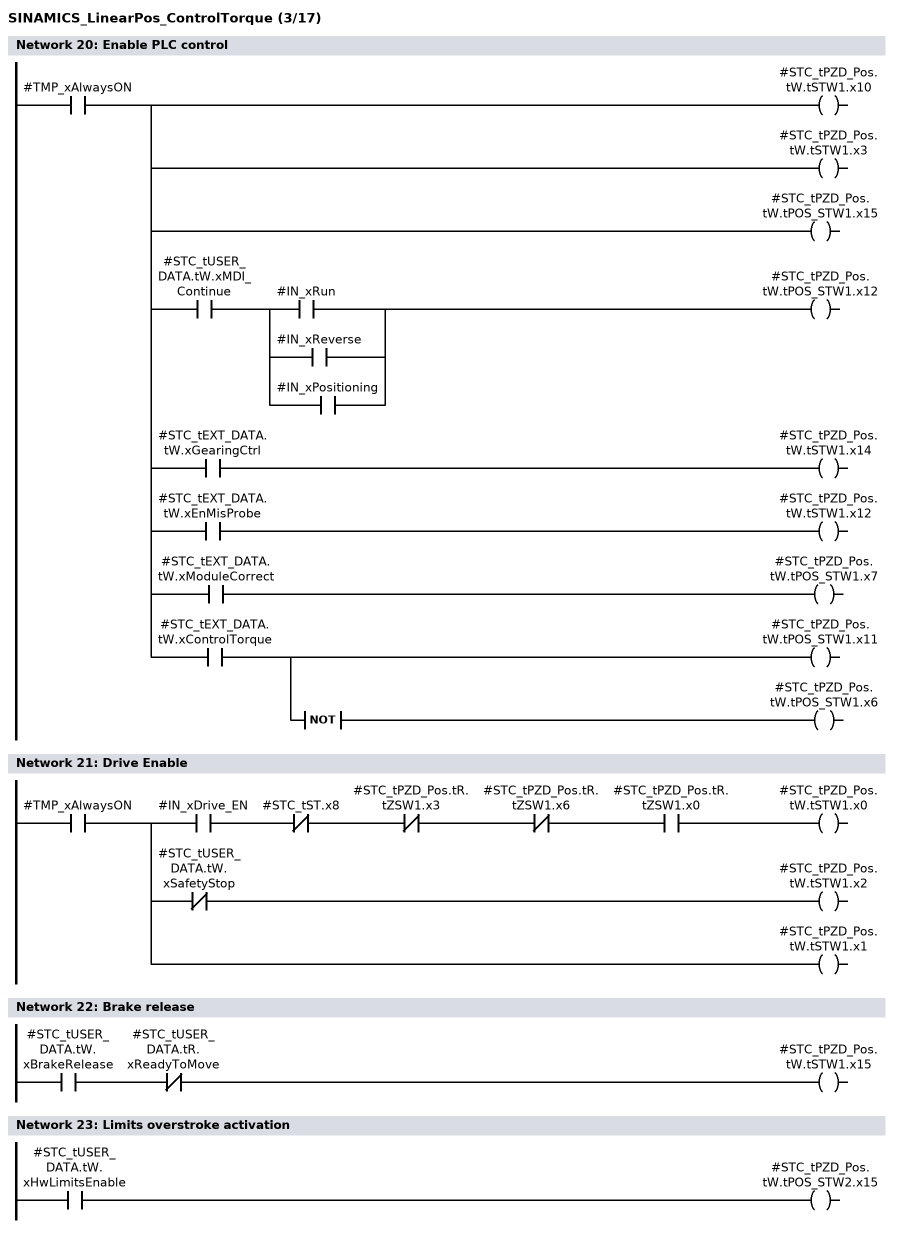
   RUNG wire#powerrail
      Contact( #TMP_xAlwaysON )
      wire#w1
      Coil( #STC_tPZD_Pos.tW.tSTW1.x10 )
   END_RUNG
   RUNG wire#w1
      Coil( #STC_tPZD_Pos.tW.tSTW1.x3 )
   END_RUNG
   RUNG wire#w1
      Coil( #STC_tPZD_Pos.tW.tPOS_STW1.x15 )
   END_RUNG
   RUNG wire#w1
      Contact( #STC_tUSER_DATA.tW.xMDI_Continue )
      wire#w2
      Contact( #IN_xRun )
      wire#w3
      Coil( #STC_tPZD_Pos.tW.tPOS_STW1.x12 )
   END_RUNG
   RUNG wire#w2
      Contact( #IN_xReverse )
   END_RUNG wire#w3
   RUNG wire#w2
      Contact( #IN_xPositioning )
   END_RUNG wire#w3
   RUNG wire#w1
      Contact( #STC_tEXT_DATA.tW.xGearingCtrl )
      Coil( #STC_tPZD_Pos.tW.tSTW1.x14 )
   END_RUNG
   RUNG wire#w1
      Contact( #STC_tEXT_DATA.tW.xEnMisProbe )
      Coil( #STC_tPZD_Pos.tW.tSTW1.x12 )
   END_RUNG
   RUNG wire#w1
      Contact( #STC_tEXT_DATA.tW.xModuleCorrect )
      Coil( #STC_tPZD_Pos.tW.tPOS_STW1.x7 )
   END_RUNG
   RUNG wire#w1
      Contact( #STC_tEXT_DATA.tW.xControlTorque )
      wire#w4
      Coil( #STC_tPZD_Pos.tW.tPOS_STW1.x11 )
   END_RUNG
   RUNG wire#w4
      Not()
      Coil( #STC_tPZD_Pos.tW.tPOS_STW1.x6 )
   END_RUNG
   // the same network as SCL:
   #STC_tPZD_Pos.tW.tSTW1.x10 := #TMP_xAlwaysON;
   #STC_tPZD_Pos.tW.tSTW1.x3 := #TMP_xAlwaysON;
   #STC_tPZD_Pos.tW.tPOS_STW1.x15 := #TMP_xAlwaysON;
   #STC_tPZD_Pos.tW.tPOS_STW1.x12 := #TMP_xAlwaysON AND #STC_tUSER_DATA.tW.xMDI_Continue AND (#IN_xRun OR #IN_xReverse OR #IN_xPositioning);
   #STC_tPZD_Pos.tW.tSTW1.x14 := #TMP_xAlwaysON AND #STC_tEXT_DATA.tW.xGearingCtrl;
   #STC_tPZD_Pos.tW.tSTW1.x12 := #TMP_xAlwaysON AND #STC_tEXT_DATA.tW.xEnMisProbe;
   #STC_tPZD_Pos.tW.tPOS_STW1.x7 := #TMP_xAlwaysON AND #STC_tEXT_DATA.tW.xModuleCorrect;
   #STC_tPZD_Pos.tW.tPOS_STW1.x11 := #TMP_xAlwaysON AND #STC_tEXT_DATA.tW.xControlTorque;
   #STC_tPZD_Pos.tW.tPOS_STW1.x6 := NOT #STC_tPZD_Pos.tW.tPOS_STW1.x11;
END_REGION

REGION Network 21: Drive Enable
   RUNG wire#powerrail
      Contact( #TMP_xAlwaysON )
      wire#w1
      Contact( #IN_xDrive_EN )
      I_Contact( #STC_tST.x8 )
      I_Contact( #STC_tPZD_Pos.tR.tZSW1.x3 )
      I_Contact( #STC_tPZD_Pos.tR.tZSW1.x6 )
      Contact( #STC_tPZD_Pos.tR.tZSW1.x0 )
      Coil( #STC_tPZD_Pos.tW.tSTW1.x0 )
   END_RUNG
   RUNG wire#w1
      I_Contact( #STC_tUSER_DATA.tW.xSafetyStop )
      Coil( #STC_tPZD_Pos.tW.tSTW1.x2 )
   END_RUNG
   RUNG wire#w1
      Coil( #STC_tPZD_Pos.tW.tSTW1.x1 )
   END_RUNG
   // the same network as SCL:
   #STC_tPZD_Pos.tW.tSTW1.x0 := #TMP_xAlwaysON AND #IN_xDrive_EN AND NOT #STC_tST.x8 AND NOT #STC_tPZD_Pos.tR.tZSW1.x3 AND NOT #STC_tPZD_Pos.tR.tZSW1.x6 AND #STC_tPZD_Pos.tR.tZSW1.x0;
   #STC_tPZD_Pos.tW.tSTW1.x2 := #TMP_xAlwaysON AND NOT #STC_tUSER_DATA.tW.xSafetyStop;
   #STC_tPZD_Pos.tW.tSTW1.x1 := #TMP_xAlwaysON;
END_REGION

REGION Network 22: Brake release
   RUNG wire#powerrail
      Contact( #STC_tUSER_DATA.tW.xBrakeRelease )
      I_Contact( #STC_tUSER_DATA.tR.xReadyToMove )
      Coil( #STC_tPZD_Pos.tW.tSTW1.x15 )
   END_RUNG
   // the same network as SCL:
   #STC_tPZD_Pos.tW.tSTW1.x15 := #STC_tUSER_DATA.tW.xBrakeRelease AND NOT #STC_tUSER_DATA.tR.xReadyToMove;
END_REGION

REGION Network 23: Limits overstroke activation
   RUNG wire#powerrail
      Contact( #STC_tUSER_DATA.tW.xHwLimitsEnable )
      Coil( #STC_tPZD_Pos.tW.tPOS_STW2.x15 )
   END_RUNG
   // the same network as SCL:
   #STC_tPZD_Pos.tW.tPOS_STW2.x15 := #STC_tUSER_DATA.tW.xHwLimitsEnable;
END_REGION

REGION Network 24: OS.Fly referencing active
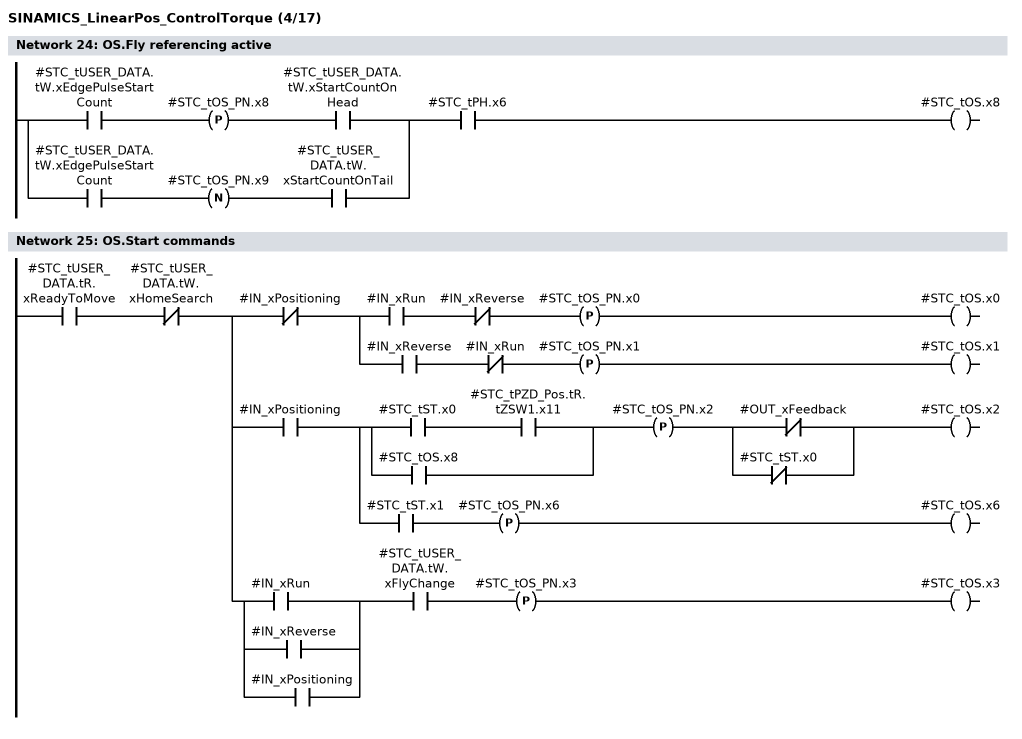
   RUNG wire#powerrail
      Contact( #STC_tUSER_DATA.tW.xEdgePulseStartCount )
      P_Trig( #STC_tOS_PN.x8 )
      Contact( #STC_tUSER_DATA.tW.xStartCountOnHead )
      wire#w1
      Contact( #STC_tPH.x6 )
      Coil( #STC_tOS.x8 )
   END_RUNG
   RUNG wire#powerrail
      Contact( #STC_tUSER_DATA.tW.xEdgePulseStartCount )
      N_Trig( #STC_tOS_PN.x9 )
      Contact( #STC_tUSER_DATA.tW.xStartCountOnTail )
   END_RUNG wire#w1
   // the same network as SCL:
   #_w1 := #STC_tUSER_DATA.tW.xEdgePulseStartCount AND NOT #STC_tOS_PN.x8;   // rising edge
   #STC_tOS_PN.x8 := #STC_tUSER_DATA.tW.xEdgePulseStartCount;
   #_w2 := NOT #STC_tUSER_DATA.tW.xEdgePulseStartCount AND #STC_tOS_PN.x9;   // falling edge
   #STC_tOS_PN.x9 := #STC_tUSER_DATA.tW.xEdgePulseStartCount;
   #STC_tOS.x8 := ((#_w1 AND #STC_tUSER_DATA.tW.xStartCountOnHead) OR (#_w2 AND #STC_tUSER_DATA.tW.xStartCountOnTail)) AND #STC_tPH.x6;
END_REGION

REGION Network 25: OS.Start commands
   RUNG wire#powerrail
      Contact( #STC_tUSER_DATA.tR.xReadyToMove )
      I_Contact( #STC_tUSER_DATA.tW.xHomeSearch )
      wire#w1
      I_Contact( #IN_xPositioning )
      wire#w2
      Contact( #IN_xRun )
      I_Contact( #IN_xReverse )
      P_Trig( #STC_tOS_PN.x0 )
      Coil( #STC_tOS.x0 )
   END_RUNG
   RUNG wire#w2
      Contact( #IN_xReverse )
      I_Contact( #IN_xRun )
      P_Trig( #STC_tOS_PN.x1 )
      Coil( #STC_tOS.x1 )
   END_RUNG
   RUNG wire#w1
      Contact( #IN_xPositioning )
      wire#w3
      Contact( #STC_tST.x0 )
      Contact( #STC_tPZD_Pos.tR.tZSW1.x11 )
      wire#w4
      P_Trig( #STC_tOS_PN.x2 )
      wire#w5
      I_Contact( #OUT_xFeedback )
      wire#w6
      Coil( #STC_tOS.x2 )
   END_RUNG
   RUNG wire#w3
      Contact( #STC_tOS.x8 )
   END_RUNG wire#w4
   RUNG wire#w5
      I_Contact( #STC_tST.x0 )
   END_RUNG wire#w6
   RUNG wire#w3
      Contact( #STC_tST.x1 )
      P_Trig( #STC_tOS_PN.x6 )
      Coil( #STC_tOS.x6 )
   END_RUNG
   RUNG wire#w1
      Contact( #IN_xRun )
      wire#w7
      Contact( #STC_tUSER_DATA.tW.xFlyChange )
      P_Trig( #STC_tOS_PN.x3 )
      Coil( #STC_tOS.x3 )
   END_RUNG
   RUNG wire#w1
      Contact( #IN_xReverse )
   END_RUNG wire#w7
   RUNG wire#w1
      Contact( #IN_xPositioning )
   END_RUNG wire#w7
   // the same network as SCL:
   #_w1 := #STC_tUSER_DATA.tR.xReadyToMove AND NOT #STC_tUSER_DATA.tW.xHomeSearch;
   #_w2 := #_w1 AND NOT #IN_xPositioning;
   #_w3 := #_w2 AND #IN_xRun AND NOT #IN_xReverse;
   #_w4 := #_w3 AND NOT #STC_tOS_PN.x0;   // rising edge
   #STC_tOS_PN.x0 := #_w3;
   #STC_tOS.x0 := #_w4;
   #_w5 := #_w2 AND #IN_xReverse AND NOT #IN_xRun;
   #_w6 := #_w5 AND NOT #STC_tOS_PN.x1;   // rising edge
   #STC_tOS_PN.x1 := #_w5;
   #STC_tOS.x1 := #_w6;
   #_w7 := #_w1 AND #IN_xPositioning;
   #_w8 := #_w7 AND ((#STC_tST.x0 AND #STC_tPZD_Pos.tR.tZSW1.x11) OR #STC_tOS.x8);
   #_w9 := #_w8 AND NOT #STC_tOS_PN.x2;   // rising edge
   #STC_tOS_PN.x2 := #_w8;
   #STC_tOS.x2 := #_w9 AND (NOT #OUT_xFeedback OR NOT #STC_tST.x0);
   #_w10 := #_w7 AND #STC_tST.x1;
   #_w11 := #_w10 AND NOT #STC_tOS_PN.x6;   // rising edge
   #STC_tOS_PN.x6 := #_w10;
   #STC_tOS.x6 := #_w11;
   #_w12 := #_w1 AND (#IN_xRun OR #IN_xReverse OR #IN_xPositioning) AND #STC_tUSER_DATA.tW.xFlyChange;
   #_w13 := #_w12 AND NOT #STC_tOS_PN.x3;   // rising edge
   #STC_tOS_PN.x3 := #_w12;
   #STC_tOS.x3 := #_w13;
END_REGION

REGION Network 26: Sending data copy
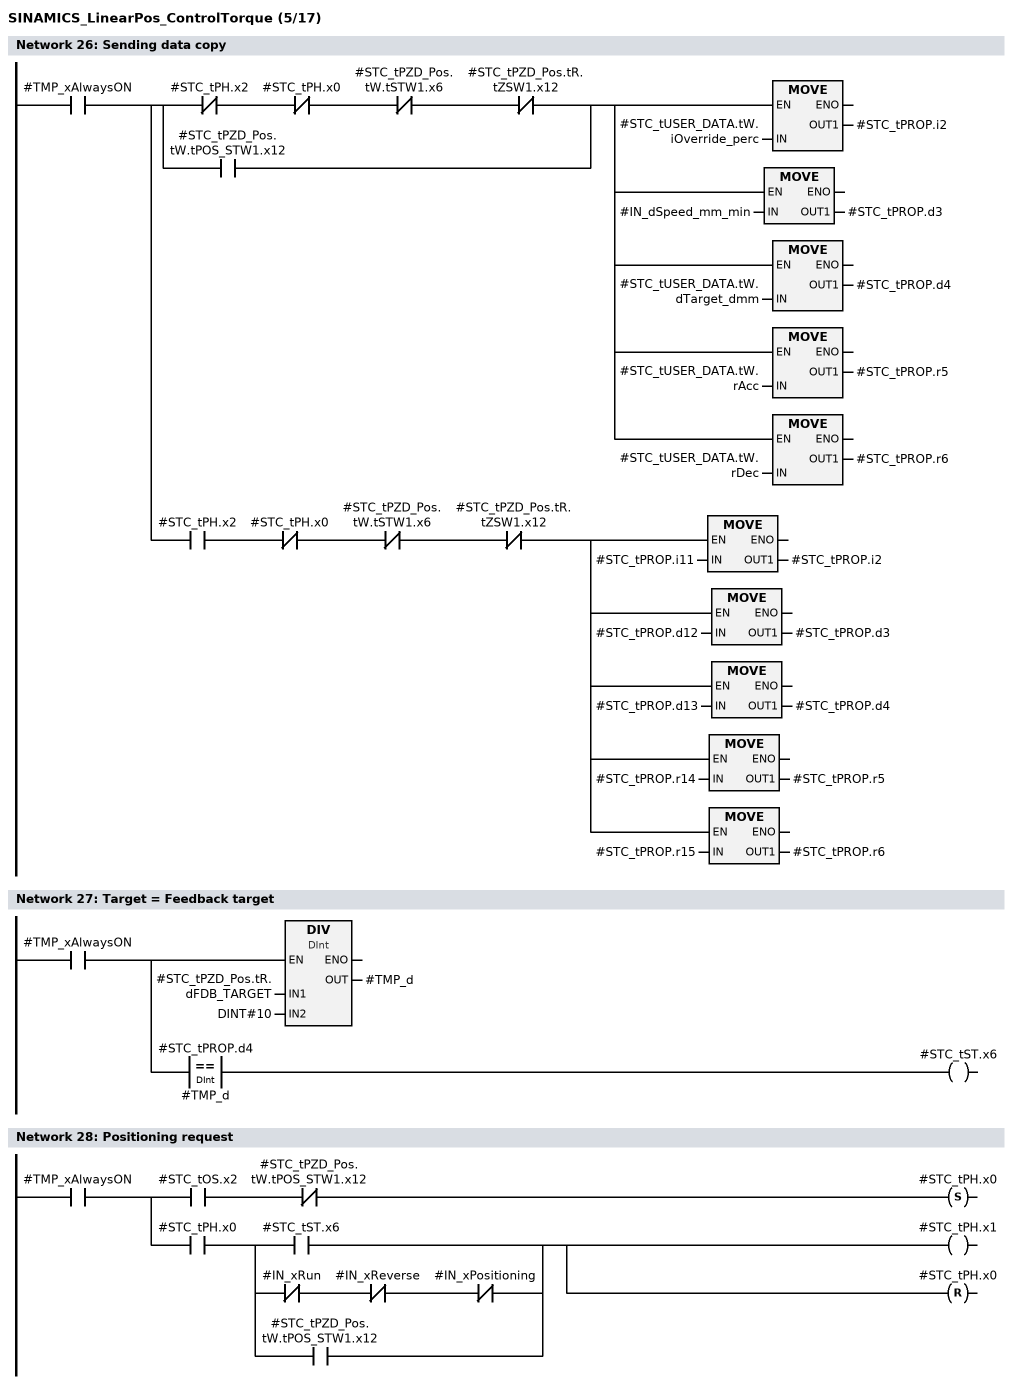
   RUNG wire#powerrail
      Contact( #TMP_xAlwaysON )
      wire#w1
      I_Contact( #STC_tPH.x2 )
      I_Contact( #STC_tPH.x0 )
      I_Contact( #STC_tPZD_Pos.tW.tSTW1.x6 )
      I_Contact( #STC_tPZD_Pos.tR.tZSW1.x12 )
      wire#w2
      { S7_GenerateENO := "TRUE" } Move(in := #STC_tUSER_DATA.tW.iOverride_perc, out1 => #STC_tPROP.i2)
   END_RUNG
   RUNG wire#w1
      Contact( #STC_tPZD_Pos.tW.tPOS_STW1.x12 )
   END_RUNG wire#w2
   RUNG wire#w2
      { S7_GenerateENO := "TRUE" } Move(in := #IN_dSpeed_mm_min, out1 => #STC_tPROP.d3)
   END_RUNG
   RUNG wire#w2
      { S7_GenerateENO := "TRUE" } Move(in := #STC_tUSER_DATA.tW.dTarget_dmm, out1 => #STC_tPROP.d4)
   END_RUNG
   RUNG wire#w2
      { S7_GenerateENO := "TRUE" } Move(in := #STC_tUSER_DATA.tW.rAcc, out1 => #STC_tPROP.r5)
   END_RUNG
   RUNG wire#w2
      { S7_GenerateENO := "TRUE" } Move(in := #STC_tUSER_DATA.tW.rDec, out1 => #STC_tPROP.r6)
   END_RUNG
   RUNG wire#w1
      Contact( #STC_tPH.x2 )
      I_Contact( #STC_tPH.x0 )
      I_Contact( #STC_tPZD_Pos.tW.tSTW1.x6 )
      I_Contact( #STC_tPZD_Pos.tR.tZSW1.x12 )
      wire#w3
      { S7_GenerateENO := "TRUE" } Move(in := #STC_tPROP.i11, out1 => #STC_tPROP.i2)
   END_RUNG
   RUNG wire#w3
      { S7_GenerateENO := "TRUE" } Move(in := #STC_tPROP.d12, out1 => #STC_tPROP.d3)
   END_RUNG
   RUNG wire#w3
      { S7_GenerateENO := "TRUE" } Move(in := #STC_tPROP.d13, out1 => #STC_tPROP.d4)
   END_RUNG
   RUNG wire#w3
      { S7_GenerateENO := "TRUE" } Move(in := #STC_tPROP.r14, out1 => #STC_tPROP.r5)
   END_RUNG
   RUNG wire#w3
      { S7_GenerateENO := "TRUE" } Move(in := #STC_tPROP.r15, out1 => #STC_tPROP.r6)
   END_RUNG
   // the same network as SCL:
   IF #TMP_xAlwaysON AND ((NOT #STC_tPH.x2 AND NOT #STC_tPH.x0 AND NOT #STC_tPZD_Pos.tW.tSTW1.x6 AND NOT #STC_tPZD_Pos.tR.tZSW1.x12) OR #STC_tPZD_Pos.tW.tPOS_STW1.x12) THEN
       #STC_tPROP.i2 := #STC_tUSER_DATA.tW.iOverride_perc;
       #STC_tPROP.d3 := #IN_dSpeed_mm_min;
       #STC_tPROP.d4 := #STC_tUSER_DATA.tW.dTarget_dmm;
       #STC_tPROP.r5 := #STC_tUSER_DATA.tW.rAcc;
       #STC_tPROP.r6 := #STC_tUSER_DATA.tW.rDec;
   END_IF;
   IF #TMP_xAlwaysON AND #STC_tPH.x2 AND NOT #STC_tPH.x0 AND NOT #STC_tPZD_Pos.tW.tSTW1.x6 AND NOT #STC_tPZD_Pos.tR.tZSW1.x12 THEN
       #STC_tPROP.i2 := #STC_tPROP.i11;
       #STC_tPROP.d3 := #STC_tPROP.d12;
       #STC_tPROP.d4 := #STC_tPROP.d13;
       #STC_tPROP.r5 := #STC_tPROP.r14;
       #STC_tPROP.r6 := #STC_tPROP.r15;
   END_IF;
END_REGION

REGION Network 27: Target = Feedback target
   RUNG wire#powerrail
      Contact( #TMP_xAlwaysON )
      wire#w1
      { S7_Templates := "SrcType := DInt"; S7_GenerateENO := "TRUE" } Div(in1 := #STC_tPZD_Pos.tR.dFDB_TARGET, in2 := DINT#10, out => #TMP_d)
   END_RUNG
   RUNG wire#w1
      { S7_Templates := "SrcType := DInt" } EQ_Contact(in1 := #STC_tPROP.d4, in2 := #TMP_d)
      Coil( #STC_tST.x6 )
   END_RUNG
   // the same network as SCL:
   IF #TMP_xAlwaysON THEN #TMP_d := #STC_tPZD_Pos.tR.dFDB_TARGET / DINT#10; END_IF;
   #STC_tST.x6 := #TMP_xAlwaysON AND (#STC_tPROP.d4 = #TMP_d);
END_REGION

REGION Network 28: Positioning request
   RUNG wire#powerrail
      Contact( #TMP_xAlwaysON )
      wire#w1
      Contact( #STC_tOS.x2 )
      I_Contact( #STC_tPZD_Pos.tW.tPOS_STW1.x12 )
      S_Coil( #STC_tPH.x0 )
   END_RUNG
   RUNG wire#w1
      Contact( #STC_tPH.x0 )
      wire#w2
      Contact( #STC_tST.x6 )
      wire#w3
      Coil( #STC_tPH.x1 )
   END_RUNG
   RUNG wire#w2
      I_Contact( #IN_xRun )
      I_Contact( #IN_xReverse )
      I_Contact( #IN_xPositioning )
   END_RUNG wire#w3
   RUNG wire#w2
      Contact( #STC_tPZD_Pos.tW.tPOS_STW1.x12 )
   END_RUNG wire#w3
   RUNG wire#w3
      R_Coil( #STC_tPH.x0 )
   END_RUNG
   // the same network as SCL:
   IF #TMP_xAlwaysON AND #STC_tOS.x2 AND NOT #STC_tPZD_Pos.tW.tPOS_STW1.x12 THEN #STC_tPH.x0 := TRUE; END_IF;
   #STC_tPH.x1 := #TMP_xAlwaysON AND #STC_tPH.x0 AND (#STC_tST.x6 OR (NOT #IN_xRun AND NOT #IN_xReverse AND NOT #IN_xPositioning) OR #STC_tPZD_Pos.tW.tPOS_STW1.x12);
   IF #STC_tPH.x1 THEN #STC_tPH.x0 := FALSE; END_IF;
END_REGION

REGION Network 29: Fly change request
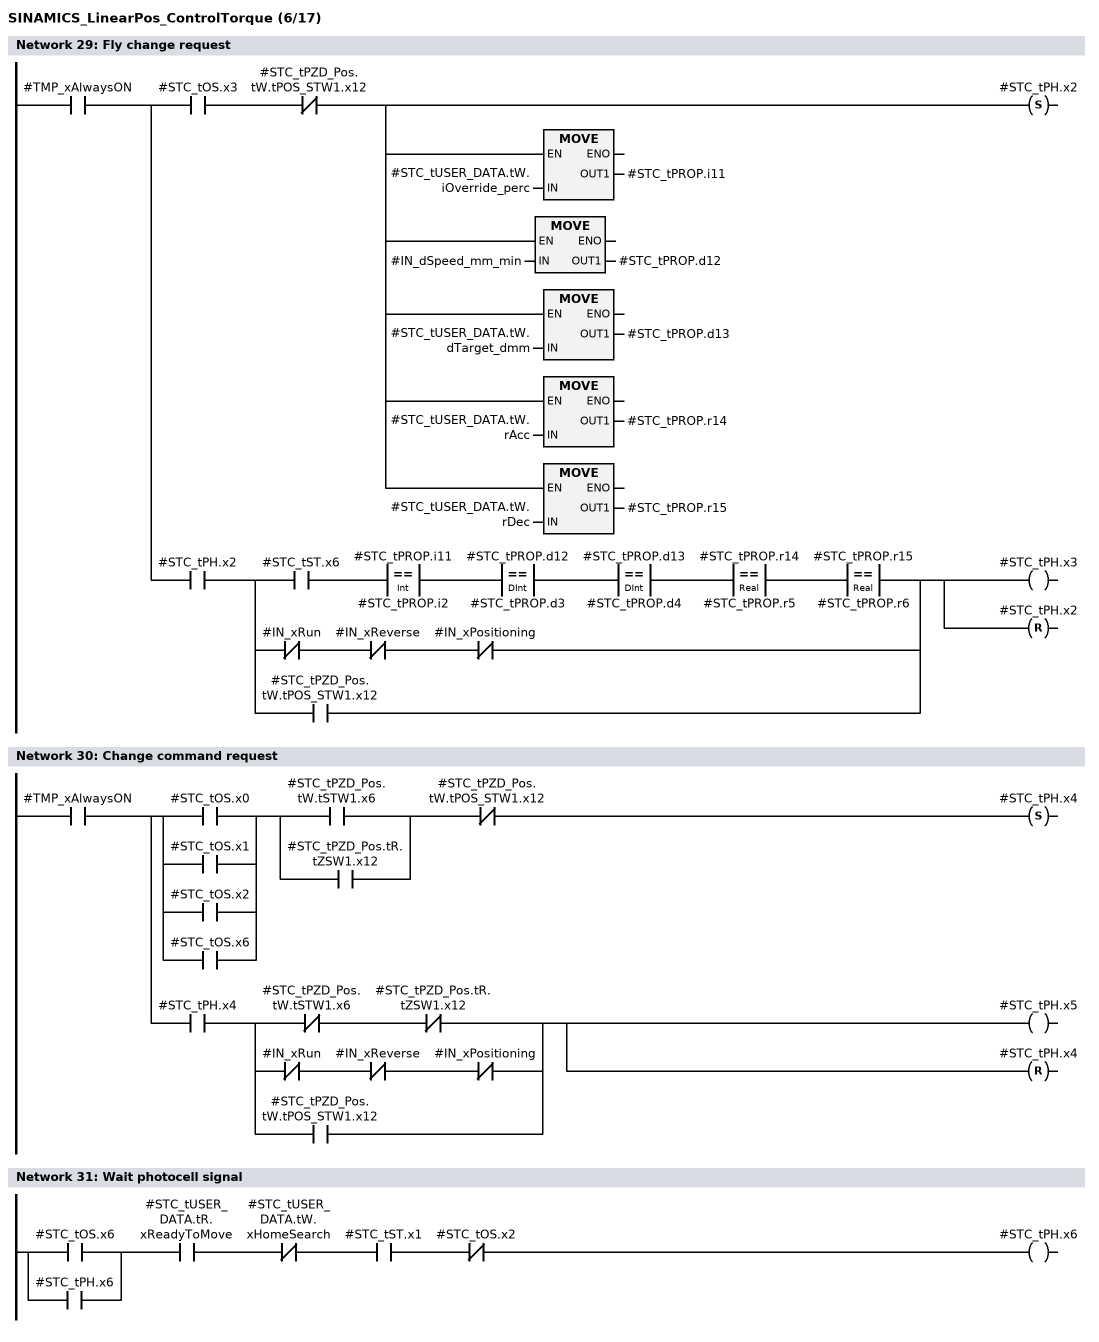
   RUNG wire#powerrail
      Contact( #TMP_xAlwaysON )
      wire#w1
      Contact( #STC_tOS.x3 )
      I_Contact( #STC_tPZD_Pos.tW.tPOS_STW1.x12 )
      wire#w2
      S_Coil( #STC_tPH.x2 )
   END_RUNG
   RUNG wire#w2
      Move(in := #STC_tUSER_DATA.tW.iOverride_perc, out1 => #STC_tPROP.i11)
   END_RUNG
   RUNG wire#w2
      Move(in := #IN_dSpeed_mm_min, out1 => #STC_tPROP.d12)
   END_RUNG
   RUNG wire#w2
      Move(in := #STC_tUSER_DATA.tW.dTarget_dmm, out1 => #STC_tPROP.d13)
   END_RUNG
   RUNG wire#w2
      Move(in := #STC_tUSER_DATA.tW.rAcc, out1 => #STC_tPROP.r14)
   END_RUNG
   RUNG wire#w2
      Move(in := #STC_tUSER_DATA.tW.rDec, out1 => #STC_tPROP.r15)
   END_RUNG
   RUNG wire#w1
      Contact( #STC_tPH.x2 )
      wire#w3
      Contact( #STC_tST.x6 )
      { S7_Templates := "SrcType := Int" } EQ_Contact(in1 := #STC_tPROP.i11, in2 := #STC_tPROP.i2)
      { S7_Templates := "SrcType := DInt" } EQ_Contact(in1 := #STC_tPROP.d12, in2 := #STC_tPROP.d3)
      { S7_Templates := "SrcType := DInt" } EQ_Contact(in1 := #STC_tPROP.d13, in2 := #STC_tPROP.d4)
      { S7_Templates := "SrcType := Real" } EQ_Contact(in1 := #STC_tPROP.r14, in2 := #STC_tPROP.r5)
      { S7_Templates := "SrcType := Real" } EQ_Contact(in1 := #STC_tPROP.r15, in2 := #STC_tPROP.r6)
      wire#w4
      Coil( #STC_tPH.x3 )
   END_RUNG
   RUNG wire#w3
      I_Contact( #IN_xRun )
      I_Contact( #IN_xReverse )
      I_Contact( #IN_xPositioning )
   END_RUNG wire#w4
   RUNG wire#w3
      Contact( #STC_tPZD_Pos.tW.tPOS_STW1.x12 )
   END_RUNG wire#w4
   RUNG wire#w4
      R_Coil( #STC_tPH.x2 )
   END_RUNG
   // the same network as SCL:
   IF #TMP_xAlwaysON AND #STC_tOS.x3 AND NOT #STC_tPZD_Pos.tW.tPOS_STW1.x12 THEN
       #STC_tPH.x2 := TRUE;
       #STC_tPROP.i11 := #STC_tUSER_DATA.tW.iOverride_perc;
       #STC_tPROP.d12 := #IN_dSpeed_mm_min;
       #STC_tPROP.d13 := #STC_tUSER_DATA.tW.dTarget_dmm;
       #STC_tPROP.r14 := #STC_tUSER_DATA.tW.rAcc;
       #STC_tPROP.r15 := #STC_tUSER_DATA.tW.rDec;
   END_IF;
   #STC_tPH.x3 := #TMP_xAlwaysON AND #STC_tPH.x2 AND ((#STC_tST.x6 AND (#STC_tPROP.i11 = #STC_tPROP.i2) AND (#STC_tPROP.d12 = #STC_tPROP.d3) AND (#STC_tPROP.d13 = #STC_tPROP.d4) AND (#STC_tPROP.r14 = #STC_tPROP.r5) AND (#STC_tPROP.r15 = #STC_tPROP.r6)) OR (NOT #IN_xRun AND NOT #IN_xReverse AND NOT #IN_xPositioning) OR #STC_tPZD_Pos.tW.tPOS_STW1.x12);
   IF #STC_tPH.x3 THEN #STC_tPH.x2 := FALSE; END_IF;
END_REGION

REGION Network 30: Change command request
   RUNG wire#powerrail
      Contact( #TMP_xAlwaysON )
      wire#w1
      Contact( #STC_tOS.x0 )
      wire#w2
      Contact( #STC_tPZD_Pos.tW.tSTW1.x6 )
      wire#w3
      I_Contact( #STC_tPZD_Pos.tW.tPOS_STW1.x12 )
      S_Coil( #STC_tPH.x4 )
   END_RUNG
   RUNG wire#w1
      Contact( #STC_tOS.x1 )
   END_RUNG wire#w2
   RUNG wire#w1
      Contact( #STC_tOS.x2 )
   END_RUNG wire#w2
   RUNG wire#w1
      Contact( #STC_tOS.x6 )
   END_RUNG wire#w2
   RUNG wire#w2
      Contact( #STC_tPZD_Pos.tR.tZSW1.x12 )
   END_RUNG wire#w3
   RUNG wire#w1
      Contact( #STC_tPH.x4 )
      wire#w4
      I_Contact( #STC_tPZD_Pos.tW.tSTW1.x6 )
      I_Contact( #STC_tPZD_Pos.tR.tZSW1.x12 )
      wire#w5
      Coil( #STC_tPH.x5 )
   END_RUNG
   RUNG wire#w4
      I_Contact( #IN_xRun )
      I_Contact( #IN_xReverse )
      I_Contact( #IN_xPositioning )
   END_RUNG wire#w5
   RUNG wire#w4
      Contact( #STC_tPZD_Pos.tW.tPOS_STW1.x12 )
   END_RUNG wire#w5
   RUNG wire#w5
      R_Coil( #STC_tPH.x4 )
   END_RUNG
   // the same network as SCL:
   IF #TMP_xAlwaysON AND (#STC_tOS.x0 OR #STC_tOS.x1 OR #STC_tOS.x2 OR #STC_tOS.x6) AND (#STC_tPZD_Pos.tW.tSTW1.x6 OR #STC_tPZD_Pos.tR.tZSW1.x12) AND NOT #STC_tPZD_Pos.tW.tPOS_STW1.x12 THEN
       #STC_tPH.x4 := TRUE;
   END_IF;
   #STC_tPH.x5 := #TMP_xAlwaysON AND #STC_tPH.x4 AND ((NOT #STC_tPZD_Pos.tW.tSTW1.x6 AND NOT #STC_tPZD_Pos.tR.tZSW1.x12) OR (NOT #IN_xRun AND NOT #IN_xReverse AND NOT #IN_xPositioning) OR #STC_tPZD_Pos.tW.tPOS_STW1.x12);
   IF #STC_tPH.x5 THEN #STC_tPH.x4 := FALSE; END_IF;
END_REGION

REGION Network 31: Wait photocell signal
   RUNG wire#powerrail
      Contact( #STC_tOS.x6 )
      wire#w1
      Contact( #STC_tUSER_DATA.tR.xReadyToMove )
      I_Contact( #STC_tUSER_DATA.tW.xHomeSearch )
      Contact( #STC_tST.x1 )
      I_Contact( #STC_tOS.x2 )
      Coil( #STC_tPH.x6 )
   END_RUNG
   RUNG wire#powerrail
      Contact( #STC_tPH.x6 )
   END_RUNG wire#w1
   // the same network as SCL:
   #STC_tPH.x6 := (#STC_tOS.x6 OR #STC_tPH.x6) AND #STC_tUSER_DATA.tR.xReadyToMove AND NOT #STC_tUSER_DATA.tW.xHomeSearch AND #STC_tST.x1 AND NOT #STC_tOS.x2;
END_REGION

REGION Network 32: Run/Reverse Commands
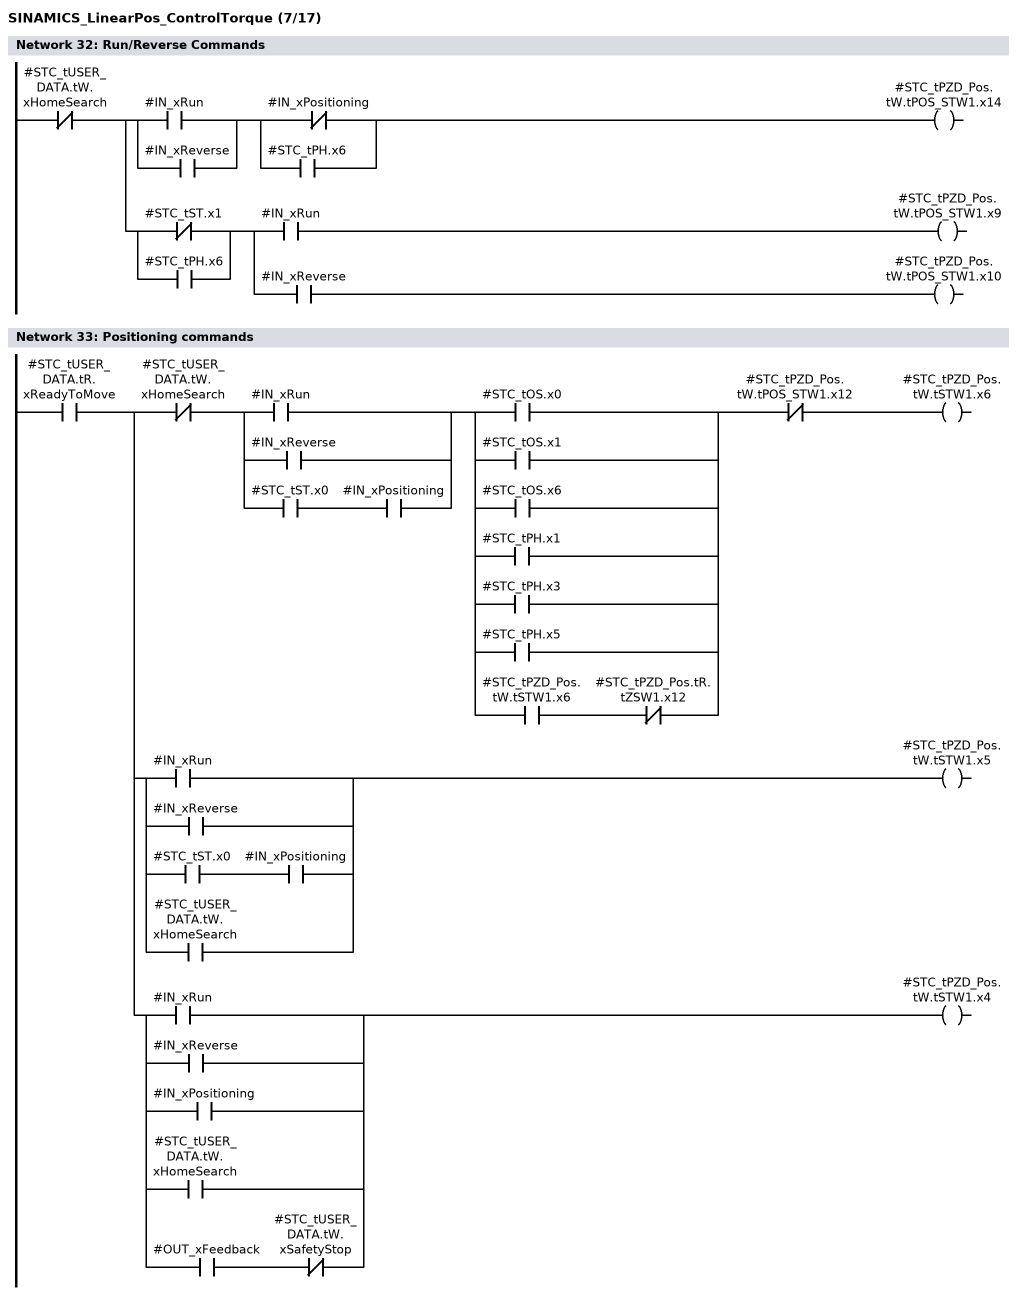
   RUNG wire#powerrail
      I_Contact( #STC_tUSER_DATA.tW.xHomeSearch )
      wire#w1
      Contact( #IN_xRun )
      wire#w2
      I_Contact( #IN_xPositioning )
      wire#w3
      Coil( #STC_tPZD_Pos.tW.tPOS_STW1.x14 )
   END_RUNG
   RUNG wire#w1
      Contact( #IN_xReverse )
   END_RUNG wire#w2
   RUNG wire#w2
      Contact( #STC_tPH.x6 )
   END_RUNG wire#w3
   RUNG wire#w1
      I_Contact( #STC_tST.x1 )
      wire#w4
      Contact( #IN_xRun )
      Coil( #STC_tPZD_Pos.tW.tPOS_STW1.x9 )
   END_RUNG
   RUNG wire#w1
      Contact( #STC_tPH.x6 )
   END_RUNG wire#w4
   RUNG wire#w4
      Contact( #IN_xReverse )
      Coil( #STC_tPZD_Pos.tW.tPOS_STW1.x10 )
   END_RUNG
   // the same network as SCL:
   #_w1 := NOT #STC_tUSER_DATA.tW.xHomeSearch;
   #STC_tPZD_Pos.tW.tPOS_STW1.x14 := #_w1 AND (#IN_xRun OR #IN_xReverse) AND (NOT #IN_xPositioning OR #STC_tPH.x6);
   #_w2 := #_w1 AND (NOT #STC_tST.x1 OR #STC_tPH.x6);
   #STC_tPZD_Pos.tW.tPOS_STW1.x9 := #_w2 AND #IN_xRun;
   #STC_tPZD_Pos.tW.tPOS_STW1.x10 := #_w2 AND #IN_xReverse;
END_REGION

REGION Network 33: Positioning commands
   RUNG wire#powerrail
      Contact( #STC_tUSER_DATA.tR.xReadyToMove )
      wire#w1
      I_Contact( #STC_tUSER_DATA.tW.xHomeSearch )
      wire#w2
      Contact( #IN_xRun )
      wire#w3
      Contact( #STC_tOS.x0 )
      wire#w4
      I_Contact( #STC_tPZD_Pos.tW.tPOS_STW1.x12 )
      Coil( #STC_tPZD_Pos.tW.tSTW1.x6 )
   END_RUNG
   RUNG wire#w2
      Contact( #IN_xReverse )
   END_RUNG wire#w3
   RUNG wire#w2
      Contact( #STC_tST.x0 )
      Contact( #IN_xPositioning )
   END_RUNG wire#w3
   RUNG wire#w3
      Contact( #STC_tOS.x1 )
   END_RUNG wire#w4
   RUNG wire#w3
      Contact( #STC_tOS.x6 )
   END_RUNG wire#w4
   RUNG wire#w3
      Contact( #STC_tPH.x1 )
   END_RUNG wire#w4
   RUNG wire#w3
      Contact( #STC_tPH.x3 )
   END_RUNG wire#w4
   RUNG wire#w3
      Contact( #STC_tPH.x5 )
   END_RUNG wire#w4
   RUNG wire#w3
      Contact( #STC_tPZD_Pos.tW.tSTW1.x6 )
      I_Contact( #STC_tPZD_Pos.tR.tZSW1.x12 )
   END_RUNG wire#w4
   RUNG wire#w1
      Contact( #IN_xRun )
      wire#w5
      Coil( #STC_tPZD_Pos.tW.tSTW1.x5 )
   END_RUNG
   RUNG wire#w1
      Contact( #IN_xReverse )
   END_RUNG wire#w5
   RUNG wire#w1
      Contact( #STC_tST.x0 )
      Contact( #IN_xPositioning )
   END_RUNG wire#w5
   RUNG wire#w1
      Contact( #STC_tUSER_DATA.tW.xHomeSearch )
   END_RUNG wire#w5
   RUNG wire#w1
      Contact( #IN_xRun )
      wire#w6
      Coil( #STC_tPZD_Pos.tW.tSTW1.x4 )
   END_RUNG
   RUNG wire#w1
      Contact( #IN_xReverse )
   END_RUNG wire#w6
   RUNG wire#w1
      Contact( #IN_xPositioning )
   END_RUNG wire#w6
   RUNG wire#w1
      Contact( #STC_tUSER_DATA.tW.xHomeSearch )
   END_RUNG wire#w6
   RUNG wire#w1
      Contact( #OUT_xFeedback )
      I_Contact( #STC_tUSER_DATA.tW.xSafetyStop )
   END_RUNG wire#w6
   // the same network as SCL:
   #STC_tPZD_Pos.tW.tSTW1.x6 := #STC_tUSER_DATA.tR.xReadyToMove AND NOT #STC_tUSER_DATA.tW.xHomeSearch AND (#IN_xRun OR #IN_xReverse OR (#STC_tST.x0 AND #IN_xPositioning)) AND (#STC_tOS.x0 OR #STC_tOS.x1 OR #STC_tOS.x6 OR #STC_tPH.x1 OR #STC_tPH.x3 OR #STC_tPH.x5 OR (#STC_tPZD_Pos.tW.tSTW1.x6 AND NOT #STC_tPZD_Pos.tR.tZSW1.x12)) AND NOT #STC_tPZD_Pos.tW.tPOS_STW1.x12;
   #STC_tPZD_Pos.tW.tSTW1.x5 := #STC_tUSER_DATA.tR.xReadyToMove AND (#IN_xRun OR #IN_xReverse OR (#STC_tST.x0 AND #IN_xPositioning) OR #STC_tUSER_DATA.tW.xHomeSearch);
   #STC_tPZD_Pos.tW.tSTW1.x4 := #STC_tUSER_DATA.tR.xReadyToMove AND (#IN_xRun OR #IN_xReverse OR #IN_xPositioning OR #STC_tUSER_DATA.tW.xHomeSearch OR (#OUT_xFeedback AND NOT #STC_tUSER_DATA.tW.xSafetyStop));
END_REGION

REGION Network 34: Choose positioning type
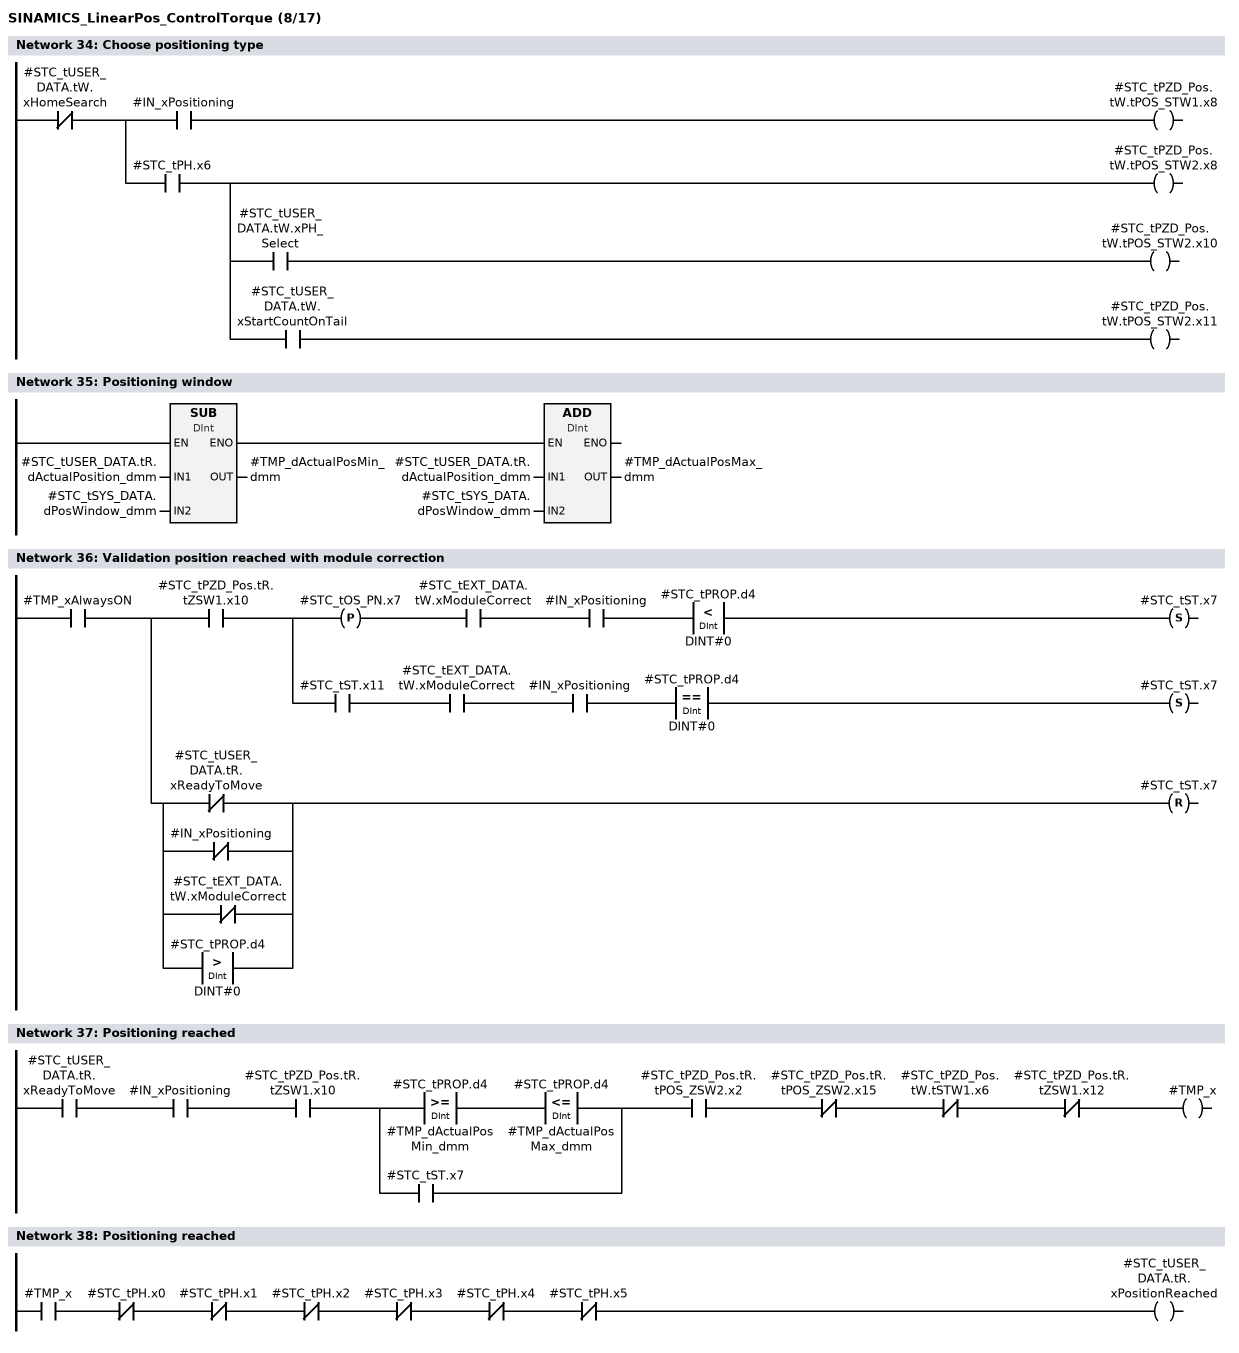
   RUNG wire#powerrail
      I_Contact( #STC_tUSER_DATA.tW.xHomeSearch )
      wire#w1
      Contact( #IN_xPositioning )
      Coil( #STC_tPZD_Pos.tW.tPOS_STW1.x8 )
   END_RUNG
   RUNG wire#w1
      Contact( #STC_tPH.x6 )
      wire#w2
      Coil( #STC_tPZD_Pos.tW.tPOS_STW2.x8 )
   END_RUNG
   RUNG wire#w2
      Contact( #STC_tUSER_DATA.tW.xPH_Select )
      Coil( #STC_tPZD_Pos.tW.tPOS_STW2.x10 )
   END_RUNG
   RUNG wire#w2
      Contact( #STC_tUSER_DATA.tW.xStartCountOnTail )
      Coil( #STC_tPZD_Pos.tW.tPOS_STW2.x11 )
   END_RUNG
   // the same network as SCL:
   #_w1 := NOT #STC_tUSER_DATA.tW.xHomeSearch;
   #STC_tPZD_Pos.tW.tPOS_STW1.x8 := #_w1 AND #IN_xPositioning;
   #STC_tPZD_Pos.tW.tPOS_STW2.x8 := #_w1 AND #STC_tPH.x6;
   #STC_tPZD_Pos.tW.tPOS_STW2.x10 := #STC_tPZD_Pos.tW.tPOS_STW2.x8 AND #STC_tUSER_DATA.tW.xPH_Select;
   #STC_tPZD_Pos.tW.tPOS_STW2.x11 := #STC_tPZD_Pos.tW.tPOS_STW2.x8 AND #STC_tUSER_DATA.tW.xStartCountOnTail;
END_REGION

REGION Network 35: Positioning window
   RUNG wire#powerrail
      { S7_Templates := "SrcType := DInt"; S7_GenerateENO := "TRUE" } Sub(in1 := #STC_tUSER_DATA.tR.dActualPosition_dmm, in2 := #STC_tSYS_DATA.dPosWindow_dmm, out => #TMP_dActualPosMin_dmm)
      { S7_Templates := "SrcType := DInt"; S7_GenerateENO := "TRUE" } Add(in1 := #STC_tUSER_DATA.tR.dActualPosition_dmm, in2 := #STC_tSYS_DATA.dPosWindow_dmm, out => #TMP_dActualPosMax_dmm)
   END_RUNG
   // the same network as SCL:
   // ENO of a box is taken as its EN; it also drops when the box reports an error
   #TMP_dActualPosMin_dmm := #STC_tUSER_DATA.tR.dActualPosition_dmm - #STC_tSYS_DATA.dPosWindow_dmm;
   #TMP_dActualPosMax_dmm := #STC_tUSER_DATA.tR.dActualPosition_dmm + #STC_tSYS_DATA.dPosWindow_dmm;
END_REGION

REGION Network 36: Validation position reached with module correction
   RUNG wire#powerrail
      Contact( #TMP_xAlwaysON )
      wire#w1
      Contact( #STC_tPZD_Pos.tR.tZSW1.x10 )
      wire#w2
      P_Trig( #STC_tOS_PN.x7 )
      Contact( #STC_tEXT_DATA.tW.xModuleCorrect )
      Contact( #IN_xPositioning )
      { S7_Templates := "SrcType := DInt" } LT_Contact(in1 := #STC_tPROP.d4, in2 := DINT#0)
      S_Coil( #STC_tST.x7 )
   END_RUNG
   RUNG wire#w2
      Contact( #STC_tST.x11 )
      Contact( #STC_tEXT_DATA.tW.xModuleCorrect )
      Contact( #IN_xPositioning )
      { S7_Templates := "SrcType := DInt" } EQ_Contact(in1 := #STC_tPROP.d4, in2 := DINT#0)
      S_Coil( #STC_tST.x7 )
   END_RUNG
   RUNG wire#w1
      I_Contact( #STC_tUSER_DATA.tR.xReadyToMove )
      wire#w3
      R_Coil( #STC_tST.x7 )
   END_RUNG
   RUNG wire#w1
      I_Contact( #IN_xPositioning )
   END_RUNG wire#w3
   RUNG wire#w1
      I_Contact( #STC_tEXT_DATA.tW.xModuleCorrect )
   END_RUNG wire#w3
   RUNG wire#w1
      { S7_Templates := "SrcType := DInt" } GT_Contact(in1 := #STC_tPROP.d4, in2 := DINT#0)
   END_RUNG wire#w3
   // the same network as SCL:
   #_w1 := #TMP_xAlwaysON AND #STC_tPZD_Pos.tR.tZSW1.x10;
   #_w2 := #_w1 AND NOT #STC_tOS_PN.x7;   // rising edge
   #STC_tOS_PN.x7 := #_w1;
   IF #_w2 AND #STC_tEXT_DATA.tW.xModuleCorrect AND #IN_xPositioning AND (#STC_tPROP.d4 < DINT#0) THEN
       #STC_tST.x7 := TRUE;
   END_IF;
   IF #_w1 AND #STC_tST.x11 AND #STC_tEXT_DATA.tW.xModuleCorrect AND #IN_xPositioning AND (#STC_tPROP.d4 = DINT#0) THEN
       #STC_tST.x7 := TRUE;
   END_IF;
   IF #TMP_xAlwaysON AND (NOT #STC_tUSER_DATA.tR.xReadyToMove OR NOT #IN_xPositioning OR NOT #STC_tEXT_DATA.tW.xModuleCorrect OR (#STC_tPROP.d4 > DINT#0)) THEN
       #STC_tST.x7 := FALSE;
   END_IF;
END_REGION

REGION Network 37: Positioning reached
   RUNG wire#powerrail
      Contact( #STC_tUSER_DATA.tR.xReadyToMove )
      Contact( #IN_xPositioning )
      Contact( #STC_tPZD_Pos.tR.tZSW1.x10 )
      wire#w1
      { S7_Templates := "SrcType := DInt" } GE_Contact(in1 := #STC_tPROP.d4, in2 := #TMP_dActualPosMin_dmm)
      { S7_Templates := "SrcType := DInt" } LE_Contact(in1 := #STC_tPROP.d4, in2 := #TMP_dActualPosMax_dmm)
      wire#w2
      Contact( #STC_tPZD_Pos.tR.tPOS_ZSW2.x2 )
      I_Contact( #STC_tPZD_Pos.tR.tPOS_ZSW2.x15 )
      I_Contact( #STC_tPZD_Pos.tW.tSTW1.x6 )
      I_Contact( #STC_tPZD_Pos.tR.tZSW1.x12 )
      Coil( #TMP_x )
   END_RUNG
   RUNG wire#w1
      Contact( #STC_tST.x7 )
   END_RUNG wire#w2
   // the same network as SCL:
   #TMP_x := #STC_tUSER_DATA.tR.xReadyToMove AND #IN_xPositioning AND #STC_tPZD_Pos.tR.tZSW1.x10 AND (((#STC_tPROP.d4 >= #TMP_dActualPosMin_dmm) AND (#STC_tPROP.d4 <= #TMP_dActualPosMax_dmm)) OR #STC_tST.x7) AND #STC_tPZD_Pos.tR.tPOS_ZSW2.x2 AND NOT #STC_tPZD_Pos.tR.tPOS_ZSW2.x15 AND NOT #STC_tPZD_Pos.tW.tSTW1.x6 AND NOT #STC_tPZD_Pos.tR.tZSW1.x12;
END_REGION

REGION Network 38: Positioning reached
   RUNG wire#powerrail
      Contact( #TMP_x )
      I_Contact( #STC_tPH.x0 )
      I_Contact( #STC_tPH.x1 )
      I_Contact( #STC_tPH.x2 )
      I_Contact( #STC_tPH.x3 )
      I_Contact( #STC_tPH.x4 )
      I_Contact( #STC_tPH.x5 )
      Coil( #STC_tUSER_DATA.tR.xPositionReached )
   END_RUNG
   // the same network as SCL:
   #STC_tUSER_DATA.tR.xPositionReached := #TMP_x AND NOT #STC_tPH.x0 AND NOT #STC_tPH.x1 AND NOT #STC_tPH.x2 AND NOT #STC_tPH.x3 AND NOT #STC_tPH.x4 AND NOT #STC_tPH.x5;
END_REGION

REGION Network 39: #####_HOMING_CYCLE_#####
END_REGION

REGION Network 40 (STL): Send homing preset
         A     #STC_tUSER_DATA.tW.xHomeSearch;
         AN    #STC_tPZD_Pos.tW.tSTW1.x11;
         JCN   PrH0;
         =     #STC_tW_MngSysReg.tST.xWrite_Request;

         L     #STC_tSYS_DATA.iPosPZD_MM;
         SLW   8;
         L     W#16#2;
         OW;
         T     #STC_tW_MngSysReg.tDATA.wRequest_refere_RequestID;
         L     #STC_tSYS_DATA.iPosPZD_MM;
         SLW   8;
         L     W#16#1;
         OW;
         T     #STC_tW_MngSysReg.tDATA.wAxis_NoOfParameters;
         L     W#16#1001;
         T     #STC_tW_MngSysReg.tDATA.wAttribute_NoOfElements;
         L     2599;
         T     #STC_tW_MngSysReg.tDATA.iParameter_number;
         L     W#16#0;
         T     #STC_tW_MngSysReg.tDATA.wSubindex;
         L     W#16#4301;
         T     #STC_tW_MngSysReg.tDATA.wFormat_NoOfValue;
         L     #STC_tSYS_DATA.iDiagAddress;
         T     #STC_tW_MngSysReg.tST.ID;
         L     47;
         T     #STC_tW_MngSysReg.tST.dINDEX;
         L     16;
         T     #STC_tW_MngSysReg.tST.uiLEN;

         L     #STC_tUSER_DATA.tW.dPreset_dmm;
         L     DINT#10;
         *D;
         T     #STC_tW_MngSysReg.tDATA.dwRegisterValue;

         CALL  #STC_tWriteRecord
         ( REQ    := #STC_tW_MngSysReg.tST.xWrite_Request,
           ID     := #STC_tW_MngSysReg.tST.ID,
           INDEX  := #STC_tW_MngSysReg.tST.dINDEX,
           LEN    := #STC_tW_MngSysReg.tST.uiLEN,
           DONE   := #STC_tW_MngSysReg.tST.xDone,
           BUSY   := #STC_tW_MngSysReg.tST.xBusy,
           ERROR  := #STC_tW_MngSysReg.tST.xError,
           STATUS := #STC_tW_MngSysReg.tST.dwSTATUS,
           RECORD := #STC_tW_MngSysReg.tDATA
         );
   PrH0: NOP   0;
END_REGION

REGION Network 41 (STL): Error during Send homing preset
         A     #STC_tW_MngSysReg.tST.xError;
         L     34;
         JC    Err;
END_REGION

REGION Network 42: Homing cycle